AUTHOR : Simatic
FAMILY : IEC
NAME : IEC_TMR
VERSION : 1.0
"IEC_TIMER"
BEGIN
END_DATA_BLOCK

DATA_BLOCK "C09_Heartbeat_Off_Timer"   // DB69
{ S7_Optimized_Access := 'TRUE' }
AUTHOR : Simatic
FAMILY : IEC
NAME : IEC_TMR
VERSION : 1.0
"IEC_TIMER"
BEGIN
END_DATA_BLOCK

DATA_BLOCK "C10_Heartbeat_On_Timer"   // DB70
{ S7_Optimized_Access := 'TRUE' }
AUTHOR : Simatic
FAMILY : IEC
NAME : IEC_TMR
VERSION : 1.0
"IEC_TIMER"
BEGIN
END_DATA_BLOCK

DATA_BLOCK "C10_Heartbeat_Off_Timer"   // DB71
{ S7_Optimized_Access := 'TRUE' }
AUTHOR : Simatic
FAMILY : IEC
NAME : IEC_TMR
VERSION : 1.0
"IEC_TIMER"
BEGIN
END_DATA_BLOCK

DATA_BLOCK "C31_Heartbeat_On_Timer"   // DB72
{ S7_Optimized_Access := 'TRUE' }
AUTHOR : Simatic
FAMILY : IEC
NAME : IEC_TMR
VERSION : 1.0
"IEC_TIMER"
BEGIN
END_DATA_BLOCK

DATA_BLOCK "C31_Heartbeat_Off_Timer"   // DB73
{ S7_Optimized_Access := 'TRUE' }
AUTHOR : Simatic
FAMILY : IEC
NAME : IEC_TMR
VERSION : 1.0
"IEC_TIMER"
BEGIN
END_DATA_BLOCK

DATA_BLOCK "C32_Heartbeat_On_Timer"   // DB74
{ S7_Optimized_Access := 'TRUE' }
AUTHOR : Simatic
FAMILY : IEC
NAME : IEC_TMR
VERSION : 1.0
"IEC_TIMER"
BEGIN
END_DATA_BLOCK

DATA_BLOCK "C32_Heartbeat_Off_Timer"   // DB75
{ S7_Optimized_Access := 'TRUE' }
AUTHOR : Simatic
FAMILY : IEC
NAME : IEC_TMR
VERSION : 1.0
"IEC_TIMER"
BEGIN
END_DATA_BLOCK

DATA_BLOCK "C33_Heartbeat_On_Timer"   // DB76
{ S7_Optimized_Access := 'TRUE' }
AUTHOR : Simatic
FAMILY : IEC
NAME : IEC_TMR
VERSION : 1.0
"IEC_TIMER"
BEGIN
END_DATA_BLOCK

DATA_BLOCK "C33_Heartbeat_Off_Timer"   // DB77
{ S7_Optimized_Access := 'TRUE' }
AUTHOR : Simatic
FAMILY : IEC
NAME : IEC_TMR
VERSION : 1.0
"IEC_TIMER"
BEGIN
END_DATA_BLOCK

DATA_BLOCK "C34_Heartbeat_On_Timer"   // DB78
{ S7_Optimized_Access := 'TRUE' }
AUTHOR : Simatic
FAMILY : IEC
NAME : IEC_TMR
VERSION : 1.0
"IEC_TIMER"
BEGIN
END_DATA_BLOCK

DATA_BLOCK "C34_Heartbeat_Off_Timer"   // DB79
{ S7_Optimized_Access := 'TRUE' }
AUTHOR : Simatic
FAMILY : IEC
NAME : IEC_TMR
VERSION : 1.0
"IEC_TIMER"
BEGIN
END_DATA_BLOCK

DATA_BLOCK "C35_Heartbeat_On_Timer"   // DB80
{ S7_Optimized_Access := 'TRUE' }
AUTHOR : Simatic
FAMILY : IEC
NAME : IEC_TMR
VERSION : 1.0
"IEC_TIMER"
BEGIN
END_DATA_BLOCK

DATA_BLOCK "C35_Heartbeat_Off_Timer"   // DB81
{ S7_Optimized_Access := 'TRUE' }
AUTHOR : Simatic
FAMILY : IEC
NAME : IEC_TMR
VERSION : 1.0
"IEC_TIMER"
BEGIN
END_DATA_BLOCK

DATA_BLOCK "C36_Heartbeat_On_Timer"   // DB82
{ S7_Optimized_Access := 'TRUE' }
AUTHOR : Simatic
FAMILY : IEC
NAME : IEC_TMR
VERSION : 1.0
"IEC_TIMER"
BEGIN
END_DATA_BLOCK

DATA_BLOCK "C36_Heartbeat_Off_Timer"   // DB83
{ S7_Optimized_Access := 'TRUE' }
AUTHOR : Simatic
FAMILY : IEC
NAME : IEC_TMR
VERSION : 1.0
"IEC_TIMER"
BEGIN
END_DATA_BLOCK

DATA_BLOCK "C37_Heartbeat_On_Timer"   // DB84
{ S7_Optimized_Access := 'TRUE' }
AUTHOR : Simatic
FAMILY : IEC
NAME : IEC_TMR
VERSION : 1.0
"IEC_TIMER"
BEGIN
END_DATA_BLOCK

DATA_BLOCK "C37_Heartbeat_Off_Timer"   // DB85
{ S7_Optimized_Access := 'TRUE' }
AUTHOR : Simatic
FAMILY : IEC
NAME : IEC_TMR
VERSION : 1.0
"IEC_TIMER"
BEGIN
END_DATA_BLOCK

DATA_BLOCK "C38_Heartbeat_On_Timer"   // DB86
{ S7_Optimized_Access := 'TRUE' }
AUTHOR : Simatic
FAMILY : IEC
NAME : IEC_TMR
VERSION : 1.0
"IEC_TIMER"
BEGIN
END_DATA_BLOCK

DATA_BLOCK "C38_Heartbeat_Off_Timer"   // DB87
{ S7_Optimized_Access := 'TRUE' }
AUTHOR : Simatic
FAMILY : IEC
NAME : IEC_TMR
VERSION : 1.0
"IEC_TIMER"
BEGIN
END_DATA_BLOCK

DATA_BLOCK "C39_Heartbeat_On_Timer"   // DB88
{ S7_Optimized_Access := 'TRUE' }
AUTHOR : Simatic
FAMILY : IEC
NAME : IEC_TMR
VERSION : 1.0
"IEC_TIMER"
BEGIN
END_DATA_BLOCK

DATA_BLOCK "C39_Heartbeat_Off_Timer"   // DB89
{ S7_Optimized_Access := 'TRUE' }
AUTHOR : Simatic
FAMILY : IEC
NAME : IEC_TMR
VERSION : 1.0
"IEC_TIMER"
BEGIN
END_DATA_BLOCK

DATA_BLOCK "C40_Heartbeat_On_Timer"   // DB90
{ S7_Optimized_Access := 'TRUE' }
AUTHOR : Simatic
FAMILY : IEC
NAME : IEC_TMR
VERSION : 1.0
"IEC_TIMER"
BEGIN
END_DATA_BLOCK

DATA_BLOCK "C40_Heartbeat_Off_Timer"   // DB91
{ S7_Optimized_Access := 'TRUE' }
AUTHOR : Simatic
FAMILY : IEC
NAME : IEC_TMR
VERSION : 1.0
"IEC_TIMER"
BEGIN
END_DATA_BLOCK

DATA_BLOCK "C41_Heartbeat_On_Timer"   // DB92
{ S7_Optimized_Access := 'TRUE' }
AUTHOR : Simatic
FAMILY : IEC
NAME : IEC_TMR
VERSION : 1.0
"IEC_TIMER"
BEGIN
END_DATA_BLOCK

DATA_BLOCK "C41_Heartbeat_Off_Timer"   // DB93
{ S7_Optimized_Access := 'TRUE' }
AUTHOR : Simatic
FAMILY : IEC
NAME : IEC_TMR
VERSION : 1.0
"IEC_TIMER"
BEGIN
END_DATA_BLOCK

DATA_BLOCK "C42_Heartbeat_On_Timer"   // DB94
{ S7_Optimized_Access := 'TRUE' }
AUTHOR : Simatic
FAMILY : IEC
NAME : IEC_TMR
VERSION : 1.0
"IEC_TIMER"
BEGIN
END_DATA_BLOCK

DATA_BLOCK "C42_Heartbeat_Off_Timer"   // DB95
{ S7_Optimized_Access := 'TRUE' }
AUTHOR : Simatic
FAMILY : IEC
NAME : IEC_TMR
VERSION : 1.0
"IEC_TIMER"
BEGIN
END_DATA_BLOCK

DATA_BLOCK "C43_Heartbeat_On_Timer"   // DB96
{ S7_Optimized_Access := 'TRUE' }
AUTHOR : Simatic
FAMILY : IEC
NAME : IEC_TMR
VERSION : 1.0
"IEC_TIMER"
BEGIN
END_DATA_BLOCK

DATA_BLOCK "C43_Heartbeat_Off_Timer"   // DB97
{ S7_Optimized_Access := 'TRUE' }
AUTHOR : Simatic
FAMILY : IEC
NAME : IEC_TMR
VERSION : 1.0
"IEC_TIMER"
BEGIN
END_DATA_BLOCK

DATA_BLOCK "C44_Heartbeat_On_Timer"   // DB98
{ S7_Optimized_Access := 'TRUE' }
AUTHOR : Simatic
FAMILY : IEC
NAME : IEC_TMR
VERSION : 1.0
"IEC_TIMER"
BEGIN
END_DATA_BLOCK

DATA_BLOCK "C44_Heartbeat_Off_Timer"   // DB99
{ S7_Optimized_Access := 'TRUE' }
AUTHOR : Simatic
FAMILY : IEC
NAME : IEC_TMR
VERSION : 1.0
"IEC_TIMER"
BEGIN
END_DATA_BLOCK

DATA_BLOCK "C45_Heartbeat_On_Timer"   // DB100
{ S7_Optimized_Access := 'TRUE' }
AUTHOR : Simatic
FAMILY : IEC
NAME : IEC_TMR
VERSION : 1.0
"IEC_TIMER"
BEGIN
END_DATA_BLOCK

DATA_BLOCK "C45_Heartbeat_Off_Timer"   // DB102
{ S7_Optimized_Access := 'TRUE' }
AUTHOR : Simatic
FAMILY : IEC
NAME : IEC_TMR
VERSION : 1.0
"IEC_TIMER"
BEGIN
END_DATA_BLOCK

DATA_BLOCK "C46_Heartbeat_On_Timer"   // DB103
{ S7_Optimized_Access := 'TRUE' }
AUTHOR : Simatic
FAMILY : IEC
NAME : IEC_TMR
VERSION : 1.0
"IEC_TIMER"
BEGIN
END_DATA_BLOCK

DATA_BLOCK "C46_Heartbeat_Off_Timer"   // DB104
{ S7_Optimized_Access := 'TRUE' }
AUTHOR : Simatic
FAMILY : IEC
NAME : IEC_TMR
VERSION : 1.0
"IEC_TIMER"
BEGIN
END_DATA_BLOCK

DATA_BLOCK "C47_Heartbeat_On_Timer"   // DB105
{ S7_Optimized_Access := 'TRUE' }
AUTHOR : Simatic
FAMILY : IEC
NAME : IEC_TMR
VERSION : 1.0
"IEC_TIMER"
BEGIN
END_DATA_BLOCK

DATA_BLOCK "C47_Heartbeat_Off_Timer"   // DB106
{ S7_Optimized_Access := 'TRUE' }
AUTHOR : Simatic
FAMILY : IEC
NAME : IEC_TMR
VERSION : 1.0
"IEC_TIMER"
BEGIN
END_DATA_BLOCK

DATA_BLOCK "C48_Heartbeat_On_Timer"   // DB107
{ S7_Optimized_Access := 'TRUE' }
AUTHOR : Simatic
FAMILY : IEC
NAME : IEC_TMR
VERSION : 1.0
"IEC_TIMER"
BEGIN
END_DATA_BLOCK

DATA_BLOCK "C48_Heartbeat_Off_Timer"   // DB108
{ S7_Optimized_Access := 'TRUE' }
AUTHOR : Simatic
FAMILY : IEC
NAME : IEC_TMR
VERSION : 1.0
"IEC_TIMER"
BEGIN
END_DATA_BLOCK

DATA_BLOCK "C49_Heartbeat_On_Timer"   // DB109
{ S7_Optimized_Access := 'TRUE' }
AUTHOR : Simatic
FAMILY : IEC
NAME : IEC_TMR
VERSION : 1.0
"IEC_TIMER"
BEGIN
END_DATA_BLOCK

DATA_BLOCK "C49_Heartbeat_Off_Timer"   // DB112
{ S7_Optimized_Access := 'TRUE' }
AUTHOR : Simatic
FAMILY : IEC
NAME : IEC_TMR
VERSION : 1.0
"IEC_TIMER"
BEGIN
END_DATA_BLOCK

DATA_BLOCK "C50_Heartbeat_On_Timer"   // DB113
{ S7_Optimized_Access := 'TRUE' }
AUTHOR : Simatic
FAMILY : IEC
NAME : IEC_TMR
VERSION : 1.0
"IEC_TIMER"
BEGIN
END_DATA_BLOCK

DATA_BLOCK "C50_Heartbeat_Off_Timer"   // DB114
{ S7_Optimized_Access := 'TRUE' }
AUTHOR : Simatic
FAMILY : IEC
NAME : IEC_TMR
VERSION : 1.0
"IEC_TIMER"
BEGIN
END_DATA_BLOCK

DATA_BLOCK "C51_Heartbeat_On_Timer"   // DB115
{ S7_Optimized_Access := 'TRUE' }
AUTHOR : Simatic
FAMILY : IEC
NAME : IEC_TMR
VERSION : 1.0
"IEC_TIMER"
BEGIN
END_DATA_BLOCK

DATA_BLOCK "C51_Heartbeat_Off_Timer"   // DB117
{ S7_Optimized_Access := 'TRUE' }
AUTHOR : Simatic
FAMILY : IEC
NAME : IEC_TMR
VERSION : 1.0
"IEC_TIMER"
BEGIN
END_DATA_BLOCK

DATA_BLOCK "C52_Heartbeat_On_Timer"   // DB118
{ S7_Optimized_Access := 'TRUE' }
AUTHOR : Simatic
FAMILY : IEC
NAME : IEC_TMR
VERSION : 1.0
"IEC_TIMER"
BEGIN
END_DATA_BLOCK

DATA_BLOCK "C52_Heartbeat_Off_Timer"   // DB119
{ S7_Optimized_Access := 'TRUE' }
AUTHOR : Simatic
FAMILY : IEC
NAME : IEC_TMR
VERSION : 1.0
"IEC_TIMER"
BEGIN
END_DATA_BLOCK

DATA_BLOCK "C53_Heartbeat_On_Timer"   // DB120
{ S7_Optimized_Access := 'TRUE' }
AUTHOR : Simatic
FAMILY : IEC
NAME : IEC_TMR
VERSION : 1.0
"IEC_TIMER"
BEGIN
END_DATA_BLOCK

DATA_BLOCK "C53_Heartbeat_Off_Timer"   // DB121
{ S7_Optimized_Access := 'TRUE' }
AUTHOR : Simatic
FAMILY : IEC
NAME : IEC_TMR
VERSION : 1.0
"IEC_TIMER"
BEGIN
END_DATA_BLOCK

DATA_BLOCK "C54_Heartbeat_On_Timer"   // DB122
{ S7_Optimized_Access := 'TRUE' }
AUTHOR : Simatic
FAMILY : IEC
NAME : IEC_TMR
VERSION : 1.0
"IEC_TIMER"
BEGIN
END_DATA_BLOCK

DATA_BLOCK "C54_Heartbeat_Off_Timer"   // DB123
{ S7_Optimized_Access := 'TRUE' }
AUTHOR : Simatic
FAMILY : IEC
NAME : IEC_TMR
VERSION : 1.0
"IEC_TIMER"
BEGIN
END_DATA_BLOCK

DATA_BLOCK "C55_Heartbeat_On_Timer"   // DB124
{ S7_Optimized_Access := 'TRUE' }
AUTHOR : Simatic
FAMILY : IEC
NAME : IEC_TMR
VERSION : 1.0
"IEC_TIMER"
BEGIN
END_DATA_BLOCK

DATA_BLOCK "C55_Heartbeat_Off_Timer"   // DB125
{ S7_Optimized_Access := 'TRUE' }
AUTHOR : Simatic
FAMILY : IEC
NAME : IEC_TMR
VERSION : 1.0
"IEC_TIMER"
BEGIN
END_DATA_BLOCK

DATA_BLOCK "C56_Heartbeat_On_Timer"   // DB126
{ S7_Optimized_Access := 'TRUE' }
AUTHOR : Simatic
FAMILY : IEC
NAME : IEC_TMR
VERSION : 1.0
"IEC_TIMER"
BEGIN
END_DATA_BLOCK

DATA_BLOCK "C56_Heartbeat_Off_Timer"   // DB127
{ S7_Optimized_Access := 'TRUE' }
AUTHOR : Simatic
FAMILY : IEC
NAME : IEC_TMR
VERSION : 1.0
"IEC_TIMER"
BEGIN
END_DATA_BLOCK

DATA_BLOCK "C57_Heartbeat_On_Timer"   // DB128
{ S7_Optimized_Access := 'TRUE' }
AUTHOR : Simatic
FAMILY : IEC
NAME : IEC_TMR
VERSION : 1.0
"IEC_TIMER"
BEGIN
END_DATA_BLOCK

DATA_BLOCK "C57_Heartbeat_Off_Timer"   // DB129
{ S7_Optimized_Access := 'TRUE' }
AUTHOR : Simatic
FAMILY : IEC
NAME : IEC_TMR
VERSION : 1.0
"IEC_TIMER"
BEGIN
END_DATA_BLOCK

DATA_BLOCK "C58_Heartbeat_On_Timer"   // DB130
{ S7_Optimized_Access := 'TRUE' }
AUTHOR : Simatic
FAMILY : IEC
NAME : IEC_TMR
VERSION : 1.0
"IEC_TIMER"
BEGIN
END_DATA_BLOCK

DATA_BLOCK "C58_Heartbeat_Off_Timer"   // DB131
{ S7_Optimized_Access := 'TRUE' }
AUTHOR : Simatic
FAMILY : IEC
NAME : IEC_TMR
VERSION : 1.0
"IEC_TIMER"
BEGIN
END_DATA_BLOCK

DATA_BLOCK "C59_Heartbeat_On_Timer"   // DB132
{ S7_Optimized_Access := 'TRUE' }
AUTHOR : Simatic
FAMILY : IEC
NAME : IEC_TMR
VERSION : 1.0
"IEC_TIMER"
BEGIN
END_DATA_BLOCK

DATA_BLOCK "C59_Heartbeat_Off_Timer"   // DB133
{ S7_Optimized_Access := 'TRUE' }
AUTHOR : Simatic
FAMILY : IEC
NAME : IEC_TMR
VERSION : 1.0
"IEC_TIMER"
BEGIN
END_DATA_BLOCK

DATA_BLOCK "C60_Heartbeat_On_Timer"   // DB134
{ S7_Optimized_Access := 'TRUE' }
AUTHOR : Simatic
FAMILY : IEC
NAME : IEC_TMR
VERSION : 1.0
"IEC_TIMER"
BEGIN
END_DATA_BLOCK

DATA_BLOCK "C60_Heartbeat_Off_Timer"   // DB135
{ S7_Optimized_Access := 'TRUE' }
AUTHOR : Simatic
FAMILY : IEC
NAME : IEC_TMR
VERSION : 1.0
"IEC_TIMER"
BEGIN
END_DATA_BLOCK

DATA_BLOCK "C61_Heartbeat_On_Timer"   // DB136
{ S7_Optimized_Access := 'TRUE' }
AUTHOR : Simatic
FAMILY : IEC
NAME : IEC_TMR
VERSION : 1.0
"IEC_TIMER"
BEGIN
END_DATA_BLOCK

DATA_BLOCK "C61_Heartbeat_Off_Timer"   // DB137
{ S7_Optimized_Access := 'TRUE' }
AUTHOR : Simatic
FAMILY : IEC
NAME : IEC_TMR
VERSION : 1.0
"IEC_TIMER"
BEGIN
END_DATA_BLOCK

DATA_BLOCK "C62_Heartbeat_On_Timer"   // DB138
{ S7_Optimized_Access := 'TRUE' }
AUTHOR : Simatic
FAMILY : IEC
NAME : IEC_TMR
VERSION : 1.0
"IEC_TIMER"
BEGIN
END_DATA_BLOCK

DATA_BLOCK "C62_Heartbeat_Off_Timer"   // DB139
{ S7_Optimized_Access := 'TRUE' }
AUTHOR : Simatic
FAMILY : IEC
NAME : IEC_TMR
VERSION : 1.0
"IEC_TIMER"
BEGIN
END_DATA_BLOCK

DATA_BLOCK "C63_Heartbeat_On_Timer"   // DB140
{ S7_Optimized_Access := 'TRUE' }
AUTHOR : Simatic
FAMILY : IEC
NAME : IEC_TMR
VERSION : 1.0
"IEC_TIMER"
BEGIN
END_DATA_BLOCK

DATA_BLOCK "C63_Heartbeat_Off_Timer"   // DB141
{ S7_Optimized_Access := 'TRUE' }
AUTHOR : Simatic
FAMILY : IEC
NAME : IEC_TMR
VERSION : 1.0
"IEC_TIMER"
BEGIN
END_DATA_BLOCK

DATA_BLOCK "C64_Heartbeat_On_Timer"   // DB142
{ S7_Optimized_Access := 'TRUE' }
AUTHOR : Simatic
FAMILY : IEC
NAME : IEC_TMR
VERSION : 1.0
"IEC_TIMER"
BEGIN
END_DATA_BLOCK

DATA_BLOCK "C64_Heartbeat_Off_Timer"   // DB143
{ S7_Optimized_Access := 'TRUE' }
AUTHOR : Simatic
FAMILY : IEC
NAME : IEC_TMR
VERSION : 1.0
"IEC_TIMER"
BEGIN
END_DATA_BLOCK

DATA_BLOCK "C65_Heartbeat_On_Timer"   // DB144
{ S7_Optimized_Access := 'TRUE' }
AUTHOR : Simatic
FAMILY : IEC
NAME : IEC_TMR
VERSION : 1.0
"IEC_TIMER"
BEGIN
END_DATA_BLOCK

DATA_BLOCK "C65_Heartbeat_Off_Timer"   // DB145
{ S7_Optimized_Access := 'TRUE' }
AUTHOR : Simatic
FAMILY : IEC
NAME : IEC_TMR
VERSION : 1.0
"IEC_TIMER"
BEGIN
END_DATA_BLOCK

DATA_BLOCK "C66_Heartbeat_On_Timer"   // DB146
{ S7_Optimized_Access := 'TRUE' }
AUTHOR : Simatic
FAMILY : IEC
NAME : IEC_TMR
VERSION : 1.0
"IEC_TIMER"
BEGIN
END_DATA_BLOCK

DATA_BLOCK "C66_Heartbeat_Off_Timer"   // DB147
{ S7_Optimized_Access := 'TRUE' }
AUTHOR : Simatic
FAMILY : IEC
NAME : IEC_TMR
VERSION : 1.0
"IEC_TIMER"
BEGIN
END_DATA_BLOCK

DATA_BLOCK "C67_Heartbeat_On_Timer"   // DB148
{ S7_Optimized_Access := 'TRUE' }
AUTHOR : Simatic
FAMILY : IEC
NAME : IEC_TMR
VERSION : 1.0
"IEC_TIMER"
BEGIN
END_DATA_BLOCK

DATA_BLOCK "C67_Heartbeat_Off_Timer"   // DB149
{ S7_Optimized_Access := 'TRUE' }
AUTHOR : Simatic
FAMILY : IEC
NAME : IEC_TMR
VERSION : 1.0
"IEC_TIMER"
BEGIN
END_DATA_BLOCK

DATA_BLOCK "C68_Heartbeat_On_Timer"   // DB150
{ S7_Optimized_Access := 'TRUE' }
AUTHOR : Simatic
FAMILY : IEC
NAME : IEC_TMR
VERSION : 1.0
"IEC_TIMER"
BEGIN
END_DATA_BLOCK

DATA_BLOCK "C68_Heartbeat_Off_Timer"   // DB151
{ S7_Optimized_Access := 'TRUE' }
AUTHOR : Simatic
FAMILY : IEC
NAME : IEC_TMR
VERSION : 1.0
"IEC_TIMER"
BEGIN
END_DATA_BLOCK

DATA_BLOCK "C69_Heartbeat_On_Timer"   // DB152
{ S7_Optimized_Access := 'TRUE' }
AUTHOR : Simatic
FAMILY : IEC
NAME : IEC_TMR
VERSION : 1.0
"IEC_TIMER"
BEGIN
END_DATA_BLOCK

DATA_BLOCK "C69_Heartbeat_Off_Timer"   // DB153
{ S7_Optimized_Access := 'TRUE' }
AUTHOR : Simatic
FAMILY : IEC
NAME : IEC_TMR
VERSION : 1.0
"IEC_TIMER"
BEGIN
END_DATA_BLOCK

DATA_BLOCK "C70_Heartbeat_On_Timer"   // DB154
{ S7_Optimized_Access := 'TRUE' }
AUTHOR : Simatic
FAMILY : IEC
NAME : IEC_TMR
VERSION : 1.0
"IEC_TIMER"
BEGIN
END_DATA_BLOCK

DATA_BLOCK "C70_Heartbeat_Off_Timer"   // DB155
{ S7_Optimized_Access := 'TRUE' }
AUTHOR : Simatic
FAMILY : IEC
NAME : IEC_TMR
VERSION : 1.0
"IEC_TIMER"
BEGIN
END_DATA_BLOCK

DATA_BLOCK "C71_Heartbeat_On_Timer"   // DB156
{ S7_Optimized_Access := 'TRUE' }
AUTHOR : Simatic
FAMILY : IEC
NAME : IEC_TMR
VERSION : 1.0
"IEC_TIMER"
BEGIN
END_DATA_BLOCK

DATA_BLOCK "C71_Heartbeat_Off_Timer"   // DB157
{ S7_Optimized_Access := 'TRUE' }
AUTHOR : Simatic
FAMILY : IEC
NAME : IEC_TMR
VERSION : 1.0
"IEC_TIMER"
BEGIN
END_DATA_BLOCK

DATA_BLOCK "C72_Heartbeat_On_Timer"   // DB158
{ S7_Optimized_Access := 'TRUE' }
AUTHOR : Simatic
FAMILY : IEC
NAME : IEC_TMR
VERSION : 1.0
"IEC_TIMER"
BEGIN
END_DATA_BLOCK

DATA_BLOCK "C72_Heartbeat_Off_Timer"   // DB159
{ S7_Optimized_Access := 'TRUE' }
AUTHOR : Simatic
FAMILY : IEC
NAME : IEC_TMR
VERSION : 1.0
"IEC_TIMER"
BEGIN
END_DATA_BLOCK

DATA_BLOCK "C73_Heartbeat_On_Timer"   // DB160
{ S7_Optimized_Access := 'TRUE' }
AUTHOR : Simatic
FAMILY : IEC
NAME : IEC_TMR
VERSION : 1.0
"IEC_TIMER"
BEGIN
END_DATA_BLOCK

DATA_BLOCK "C73_Heartbeat_Off_Timer"   // DB161
{ S7_Optimized_Access := 'TRUE' }
AUTHOR : Simatic
FAMILY : IEC
NAME : IEC_TMR
VERSION : 1.0
"IEC_TIMER"
BEGIN
END_DATA_BLOCK

DATA_BLOCK "C74_Heartbeat_On_Timer"   // DB162
{ S7_Optimized_Access := 'TRUE' }
AUTHOR : Simatic
FAMILY : IEC
NAME : IEC_TMR
VERSION : 1.0
"IEC_TIMER"
BEGIN
END_DATA_BLOCK

DATA_BLOCK "C74_Heartbeat_Off_Timer"   // DB163
{ S7_Optimized_Access := 'TRUE' }
AUTHOR : Simatic
FAMILY : IEC
NAME : IEC_TMR
VERSION : 1.0
"IEC_TIMER"
BEGIN
END_DATA_BLOCK

DATA_BLOCK "C75_Heartbeat_On_Timer"   // DB164
{ S7_Optimized_Access := 'TRUE' }
AUTHOR : Simatic
FAMILY : IEC
NAME : IEC_TMR
VERSION : 1.0
"IEC_TIMER"
BEGIN
END_DATA_BLOCK

DATA_BLOCK "C75_Heartbeat_Off_Timer"   // DB165
{ S7_Optimized_Access := 'TRUE' }
AUTHOR : Simatic
FAMILY : IEC
NAME : IEC_TMR
VERSION : 1.0
"IEC_TIMER"
BEGIN
END_DATA_BLOCK

DATA_BLOCK "C76_Heartbeat_On_Timer"   // DB166
{ S7_Optimized_Access := 'TRUE' }
AUTHOR : Simatic
FAMILY : IEC
NAME : IEC_TMR
VERSION : 1.0
"IEC_TIMER"
BEGIN
END_DATA_BLOCK

DATA_BLOCK "C76_Heartbeat_Off_Timer"   // DB167
{ S7_Optimized_Access := 'TRUE' }
AUTHOR : Simatic
FAMILY : IEC
NAME : IEC_TMR
VERSION : 1.0
"IEC_TIMER"
BEGIN
END_DATA_BLOCK

DATA_BLOCK "C77_Heartbeat_On_Timer"   // DB168
{ S7_Optimized_Access := 'TRUE' }
AUTHOR : Simatic
FAMILY : IEC
NAME : IEC_TMR
VERSION : 1.0
"IEC_TIMER"
BEGIN
END_DATA_BLOCK

DATA_BLOCK "C77_Heartbeat_Off_Timer"   // DB169
{ S7_Optimized_Access := 'TRUE' }
AUTHOR : Simatic
FAMILY : IEC
NAME : IEC_TMR
VERSION : 1.0
"IEC_TIMER"
BEGIN
END_DATA_BLOCK

DATA_BLOCK "C78_Heartbeat_On_Timer"   // DB170
{ S7_Optimized_Access := 'TRUE' }
AUTHOR : Simatic
FAMILY : IEC
NAME : IEC_TMR
VERSION : 1.0
"IEC_TIMER"
BEGIN
END_DATA_BLOCK

DATA_BLOCK "C78_Heartbeat_Off_Timer"   // DB171
{ S7_Optimized_Access := 'TRUE' }
AUTHOR : Simatic
FAMILY : IEC
NAME : IEC_TMR
VERSION : 1.0
"IEC_TIMER"
BEGIN
END_DATA_BLOCK

DATA_BLOCK "C79_Heartbeat_On_Timer"   // DB172
{ S7_Optimized_Access := 'TRUE' }
AUTHOR : Simatic
FAMILY : IEC
NAME : IEC_TMR
VERSION : 1.0
"IEC_TIMER"
BEGIN
END_DATA_BLOCK

DATA_BLOCK "C79_Heartbeat_Off_Timer"   // DB173
{ S7_Optimized_Access := 'TRUE' }
AUTHOR : Simatic
FAMILY : IEC
NAME : IEC_TMR
VERSION : 1.0
"IEC_TIMER"
BEGIN
END_DATA_BLOCK

DATA_BLOCK "C80_Heartbeat_On_Timer"   // DB174
{ S7_Optimized_Access := 'TRUE' }
AUTHOR : Simatic
FAMILY : IEC
NAME : IEC_TMR
VERSION : 1.0
"IEC_TIMER"
BEGIN
END_DATA_BLOCK

DATA_BLOCK "C80_Heartbeat_Off_Timer"   // DB175
{ S7_Optimized_Access := 'TRUE' }
AUTHOR : Simatic
FAMILY : IEC
NAME : IEC_TMR
VERSION : 1.0
"IEC_TIMER"
BEGIN
END_DATA_BLOCK

DATA_BLOCK "C81_Heartbeat_On_Timer"   // DB176
{ S7_Optimized_Access := 'TRUE' }
AUTHOR : Simatic
FAMILY : IEC
NAME : IEC_TMR
VERSION : 1.0
"IEC_TIMER"
BEGIN
END_DATA_BLOCK

DATA_BLOCK "C81_Heartbeat_Off_Timer"   // DB177
{ S7_Optimized_Access := 'TRUE' }
AUTHOR : Simatic
FAMILY : IEC
NAME : IEC_TMR
VERSION : 1.0
"IEC_TIMER"
BEGIN
END_DATA_BLOCK

DATA_BLOCK "C82_Heartbeat_On_Timer"   // DB178
{ S7_Optimized_Access := 'TRUE' }
AUTHOR : Simatic
FAMILY : IEC
NAME : IEC_TMR
VERSION : 1.0
"IEC_TIMER"
BEGIN
END_DATA_BLOCK

DATA_BLOCK "C82_Heartbeat_Off_Timer"   // DB179
{ S7_Optimized_Access := 'TRUE' }
AUTHOR : Simatic
FAMILY : IEC
NAME : IEC_TMR
VERSION : 1.0
"IEC_TIMER"
BEGIN
END_DATA_BLOCK

// folder: UserDiag

DATA_BLOCK "UserDiag_InstMain"   // DB2000
{ S7_Optimized_Access := 'TRUE' }
VERSION : 0.1
"UserDiag_Main"
BEGIN
END_DATA_BLOCK

DATA_BLOCK "UserDiag_DiagnosticsData"   // DB2001
TITLE = Diagosis data DB
{ S7_Optimized_Access := 'TRUE' }
VERSION : 0.1
   VAR
      plcData : "UserDiag_typePLC";   // PLC diagnostics data
      ioSystemData : Array[1.."USERDIAG_IO_SYSTEMS_UPPER_LIM"] of "UserDiag_typeIOSystem";   // IO-System diagnostics data
      startDiag : Bool := False;   // Startflag for diagnostic
   END_VAR
BEGIN
END_DATA_BLOCK

DATA_BLOCK "UserDiag_HmiData"   // DB2002
{ S7_Optimized_Access := 'TRUE' }
VERSION : 0.1
BEGIN
END_DATA_BLOCK

DATA_BLOCK "UserDiag_InstDiagnosticsStartup"   // DB2005
{ S7_Optimized_Access := 'TRUE' }
VERSION : 0.1
"UserDiag_Diagnostics"
BEGIN
END_DATA_BLOCK

// folder: (top level)

ORGANIZATION_BLOCK "SDC_Carrier_Transfer"   // OB30, LAD, CyclicInterrupt
{ S7_Optimized_Access := 'TRUE' }
VERSION : 0.1
   VAR_INPUT
      Initial_Call : Bool;   // Initial call of this OB
      Event_Count : Int;   // Events discarded
   END_VAR
BEGIN
END_ORGANIZATION_BLOCK

ORGANIZATION_BLOCK "Carrier_SDC_Transfer"   // OB31, LAD, CyclicInterrupt
{ S7_Optimized_Access := 'TRUE' }
VERSION : 0.1
   VAR_INPUT
      Initial_Call : Bool;   // Initial call of this OB
      Event_Count : Int;   // Events discarded
   END_VAR
BEGIN
END_ORGANIZATION_BLOCK

// folder: 01_OBs

ORGANIZATION_BLOCK "Main"   // OB1, LAD, ProgramCycle
TITLE = "Main Program Sweep (Cycle)"
{ S7_Optimized_Access := 'FALSE' }
VERSION : 0.1
   VAR_TEMP
      EV_CLASS : Byte;   // Bits 0-3 = 1:Coming event, Bits 4-7 = 1:Event class 1
      SCAN_1 : Byte;   // 1:Initial call of the OB, 3: Call 2-n of the OB
      PRIORITY : Byte;   // Priority of OB Execution
      OB_NUMBR : Byte;   // OB number
      RESERVED_1 : Byte;   // Reserved for system
      RESERVED_2 : Byte;   // Reserved for system
      PREV_CYCLE : Int;   // Previous program cycle time (milliseconds)
      MIN_CYCLE : Int;   // Minimum program cycle time (milliseconds)
      MAX_CYCLE : Int;   // Maximum program cycle time (milliseconds)
      DATE_TIME : Date_And_Time;   // Date and time OB started
      tempread : Bool;
      tempposition : Word;
      tempdatareceive : Word;
   END_VAR
   VAR_TEMP   // added for the SCL form of the ladder/FBD networks
      _w1 : Bool;
      _w2 : Bool;
   END_VAR
BEGIN

REGION Network 1
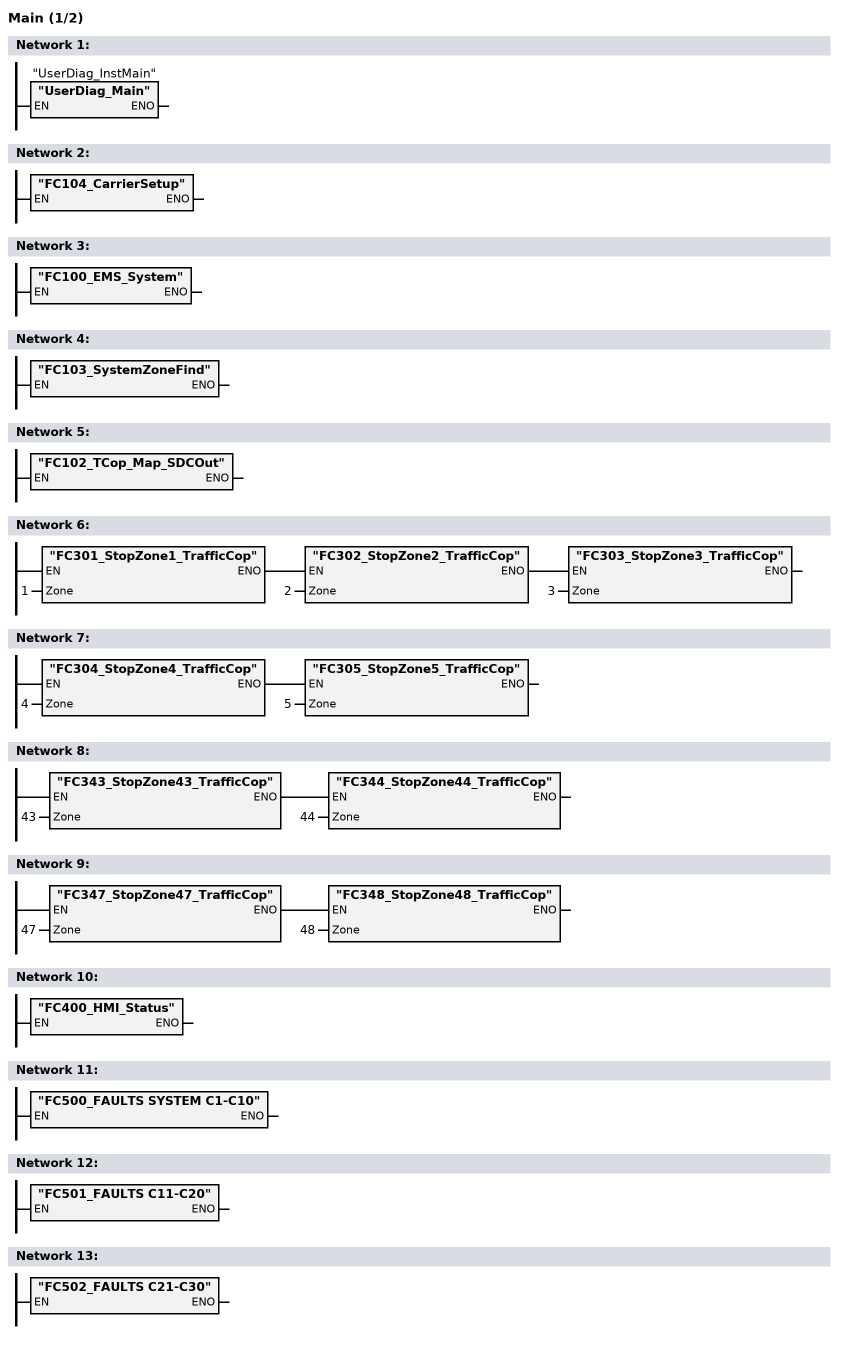
   RUNG wire#powerrail
      "UserDiag_InstMain"()
   END_RUNG
   // the same network as SCL:
   "UserDiag_InstMain"();   // "UserDiag_Main"
END_REGION

REGION Network 2
   RUNG wire#powerrail
      "FC104_CarrierSetup"()
   END_RUNG
   // the same network as SCL:
   "FC104_CarrierSetup"();
END_REGION

REGION Network 3
   RUNG wire#powerrail
      "FC100_EMS_System"()
   END_RUNG
   // the same network as SCL:
   "FC100_EMS_System"();
END_REGION

REGION Network 4
   RUNG wire#powerrail
      "FC103_SystemZoneFind"()
   END_RUNG
   // the same network as SCL:
   "FC103_SystemZoneFind"();
END_REGION

REGION Network 5
   RUNG wire#powerrail
      "FC102_TCop_Map_SDCOut"()
   END_RUNG
   // the same network as SCL:
   "FC102_TCop_Map_SDCOut"();
END_REGION

REGION Network 6
   RUNG wire#powerrail
      "FC301_StopZone1_TrafficCop"(Zone := 1)
      "FC302_StopZone2_TrafficCop"(Zone := 2)
      "FC303_StopZone3_TrafficCop"(Zone := 3)
   END_RUNG
   // the same network as SCL:
   "FC301_StopZone1_TrafficCop"(Zone := 1, ENO => #_w1);
   "FC302_StopZone2_TrafficCop"(EN := #_w1, Zone := 2, ENO => #_w2);
   IF #_w2 THEN "FC303_StopZone3_TrafficCop"(Zone := 3); END_IF;
END_REGION

REGION Network 7
   RUNG wire#powerrail
      "FC304_StopZone4_TrafficCop"(Zone := 4)
      "FC305_StopZone5_TrafficCop"(Zone := 5)
   END_RUNG
   // the same network as SCL:
   "FC304_StopZone4_TrafficCop"(Zone := 4, ENO => #_w1);
   IF #_w1 THEN "FC305_StopZone5_TrafficCop"(Zone := 5); END_IF;
END_REGION

REGION Network 8
   RUNG wire#powerrail
      "FC343_StopZone43_TrafficCop"(Zone := 43)
      "FC344_StopZone44_TrafficCop"(Zone := 44)
   END_RUNG
   // the same network as SCL:
   "FC343_StopZone43_TrafficCop"(Zone := 43, ENO => #_w1);
   IF #_w1 THEN "FC344_StopZone44_TrafficCop"(Zone := 44); END_IF;
END_REGION

REGION Network 9
   RUNG wire#powerrail
      "FC347_StopZone47_TrafficCop"(Zone := 47)
      "FC348_StopZone48_TrafficCop"(Zone := 48)
   END_RUNG
   // the same network as SCL:
   "FC347_StopZone47_TrafficCop"(Zone := 47, ENO => #_w1);
   IF #_w1 THEN "FC348_StopZone48_TrafficCop"(Zone := 48); END_IF;
END_REGION

REGION Network 10
   RUNG wire#powerrail
      "FC400_HMI_Status"()
   END_RUNG
   // the same network as SCL:
   "FC400_HMI_Status"();
END_REGION

REGION Network 11
   RUNG wire#powerrail
      "FC500_FAULTS SYSTEM C1-C10"()
   END_RUNG
   // the same network as SCL:
   "FC500_FAULTS SYSTEM C1-C10"();
END_REGION

REGION Network 12
   RUNG wire#powerrail
      "FC501_FAULTS C11-C20"()
   END_RUNG
   // the same network as SCL:
   "FC501_FAULTS C11-C20"();
END_REGION

REGION Network 13
   RUNG wire#powerrail
      "FC502_FAULTS C21-C30"()
   END_RUNG
   // the same network as SCL:
   "FC502_FAULTS C21-C30"();
END_REGION

REGION Network 14
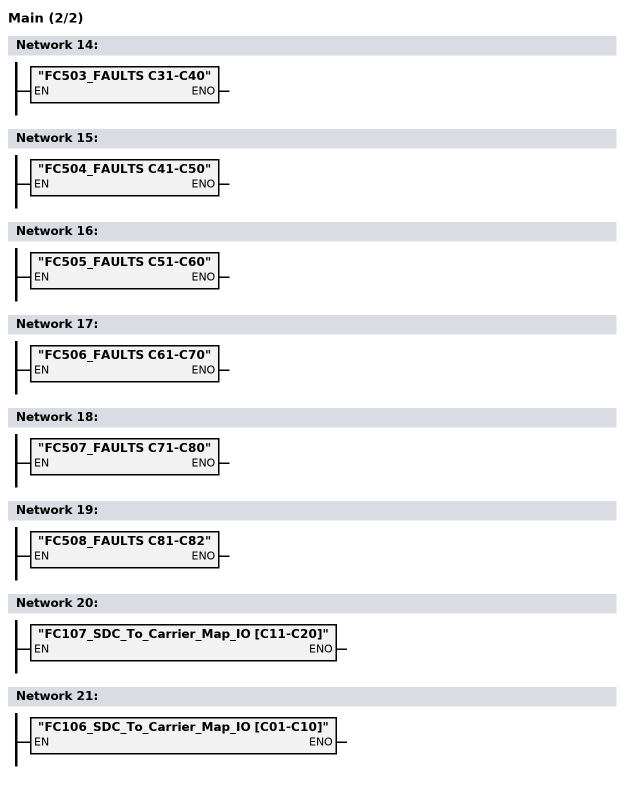
   RUNG wire#powerrail
      "FC503_FAULTS C31-C40"()
   END_RUNG
   // the same network as SCL:
   "FC503_FAULTS C31-C40"();
END_REGION

REGION Network 15
   RUNG wire#powerrail
      "FC504_FAULTS C41-C50"()
   END_RUNG
   // the same network as SCL:
   "FC504_FAULTS C41-C50"();
END_REGION

REGION Network 16
   RUNG wire#powerrail
      "FC505_FAULTS C51-C60"()
   END_RUNG
   // the same network as SCL:
   "FC505_FAULTS C51-C60"();
END_REGION

REGION Network 17
   RUNG wire#powerrail
      "FC506_FAULTS C61-C70"()
   END_RUNG
   // the same network as SCL:
   "FC506_FAULTS C61-C70"();
END_REGION

REGION Network 18
   RUNG wire#powerrail
      "FC507_FAULTS C71-C80"()
   END_RUNG
   // the same network as SCL:
   "FC507_FAULTS C71-C80"();
END_REGION

REGION Network 19
   RUNG wire#powerrail
      "FC508_FAULTS C81-C82"()
   END_RUNG
   // the same network as SCL:
   "FC508_FAULTS C81-C82"();
END_REGION

REGION Network 20
   RUNG wire#powerrail
      "FC107_SDC_To_Carrier_Map_IO [C11-C20]"()
   END_RUNG
   // the same network as SCL:
   "FC107_SDC_To_Carrier_Map_IO [C11-C20]"();
END_REGION

REGION Network 21
   RUNG wire#powerrail
      "FC106_SDC_To_Carrier_Map_IO [C01-C10]"()
   END_RUNG
   // the same network as SCL:
   "FC106_SDC_To_Carrier_Map_IO [C01-C10]"();
END_REGION
END_ORGANIZATION_BLOCK

ORGANIZATION_BLOCK "Startup"   // OB100, LAD, Startup
TITLE = "Complete Restart"
{ S7_Optimized_Access := 'TRUE' }
VERSION : 0.1
// //============================================================================
// //SIEMENS AG
// //(c)Copyright 2017 All Rights Reserved
// //-----------------------------------------------------------------------------
// //Library: -
// //Tested with: S7-1516-3 PN/DP FW 2.5
// //Engineering: TIA Portal V14 Update1
// //Restrictions: -
// //Requirements: -
// //Functionality: Startup OB for Diagnostics
// //-----------------------------------------------------------------------------
// //Change log table:
// //Version  Date              Expert in charge                               Changes applied
// //01.00.00 25.04.2017 Siemens Industry Online Support First released version
// //============================================================================
   VAR_INPUT
      LostRetentive : Bool;   // True if retentive data are lost
      LostRTC : Bool;   // True if date and time are lost
   END_VAR
   VAR_TEMP
      index : Int;
   END_VAR
BEGIN

REGION Network 1: Set start user diagnostic
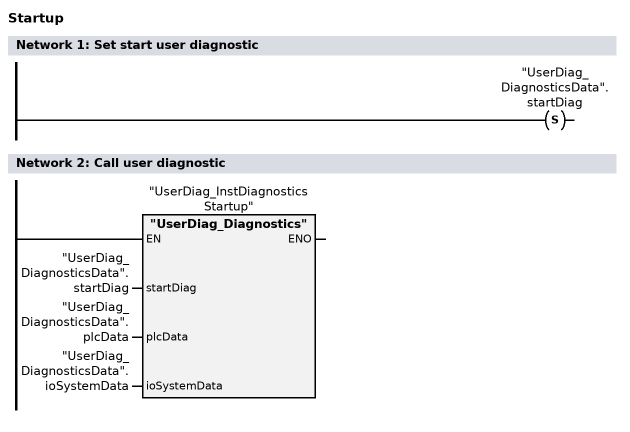
   RUNG wire#powerrail
      S_Coil( "UserDiag_DiagnosticsData".startDiag )
   END_RUNG
   // the same network as SCL:
   "UserDiag_DiagnosticsData".startDiag := TRUE;
END_REGION

REGION Network 2: Call user diagnostic
   RUNG wire#powerrail
      "UserDiag_InstDiagnosticsStartup"(startDiag := "UserDiag_DiagnosticsData".startDiag, plcData := "UserDiag_DiagnosticsData".plcData, ioSystemData := "UserDiag_DiagnosticsData".ioSystemData)
   END_RUNG
   // the same network as SCL:
   "UserDiag_InstDiagnosticsStartup"(startDiag := "UserDiag_DiagnosticsData".startDiag,   // "UserDiag_Diagnostics"
                           plcData := "UserDiag_DiagnosticsData".plcData,
                           ioSystemData := "UserDiag_DiagnosticsData".ioSystemData);
END_REGION
END_ORGANIZATION_BLOCK

ORGANIZATION_BLOCK "Cyclic SDC TO EMS"   // OB300, LAD, CyclicInterrupt
{ S7_Optimized_Access := 'TRUE' }
VERSION : 0.1
   VAR_INPUT
      Initial_Call : Bool;   // Initial call of this OB
      Event_Count : Int;   // Events discarded
   END_VAR
BEGIN
END_ORGANIZATION_BLOCK

// folder: 03_FBs

FUNCTION_BLOCK "FB110_FirstCarrierTCopMotionFB"   // FB110, LAD
{ S7_Optimized_Access := 'TRUE' }